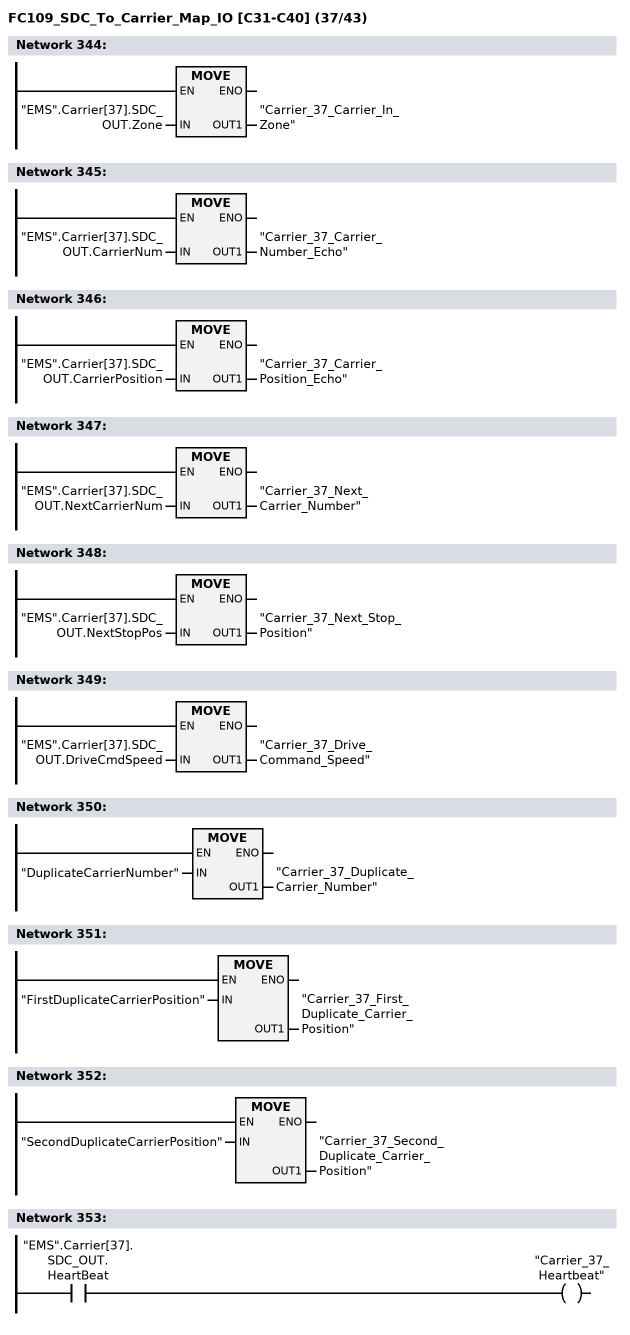
   RUNG wire#powerrail
      Move(in := "EMS".Carrier[37].SDC_OUT.Zone, out1 => "Carrier_37_Carrier_In_Zone")
   END_RUNG
   // the same network as SCL:
   "Carrier_37_Carrier_In_Zone" := "EMS".Carrier[37].SDC_OUT.Zone;
END_REGION

REGION Network 345
   RUNG wire#powerrail
      Move(in := "EMS".Carrier[37].SDC_OUT.CarrierNum, out1 => "Carrier_37_Carrier_Number_Echo")
   END_RUNG
   // the same network as SCL:
   "Carrier_37_Carrier_Number_Echo" := "EMS".Carrier[37].SDC_OUT.CarrierNum;
END_REGION

REGION Network 346
   RUNG wire#powerrail
      Move(in := "EMS".Carrier[37].SDC_OUT.CarrierPosition, out1 => "Carrier_37_Carrier_Position_Echo")
   END_RUNG
   // the same network as SCL:
   "Carrier_37_Carrier_Position_Echo" := "EMS".Carrier[37].SDC_OUT.CarrierPosition;
END_REGION

REGION Network 347
   RUNG wire#powerrail
      Move(in := "EMS".Carrier[37].SDC_OUT.NextCarrierNum, out1 => "Carrier_37_Next_Carrier_Number")
   END_RUNG
   // the same network as SCL:
   "Carrier_37_Next_Carrier_Number" := "EMS".Carrier[37].SDC_OUT.NextCarrierNum;
END_REGION

REGION Network 348
   RUNG wire#powerrail
      Move(in := "EMS".Carrier[37].SDC_OUT.NextStopPos, out1 => "Carrier_37_Next_Stop_Position")
   END_RUNG
   // the same network as SCL:
   "Carrier_37_Next_Stop_Position" := "EMS".Carrier[37].SDC_OUT.NextStopPos;
END_REGION

REGION Network 349
   RUNG wire#powerrail
      Move(in := "EMS".Carrier[37].SDC_OUT.DriveCmdSpeed, out1 => "Carrier_37_Drive_Command_Speed")
   END_RUNG
   // the same network as SCL:
   "Carrier_37_Drive_Command_Speed" := "EMS".Carrier[37].SDC_OUT.DriveCmdSpeed;
END_REGION

REGION Network 350
   RUNG wire#powerrail
      Move(in := "DuplicateCarrierNumber", out1 => "Carrier_37_Duplicate_Carrier_Number")
   END_RUNG
   // the same network as SCL:
   "Carrier_37_Duplicate_Carrier_Number" := "DuplicateCarrierNumber";
END_REGION

REGION Network 351
   RUNG wire#powerrail
      Move(in := "FirstDuplicateCarrierPosition", out1 => "Carrier_37_First_Duplicate_Carrier_Position")
   END_RUNG
   // the same network as SCL:
   "Carrier_37_First_Duplicate_Carrier_Position" := "FirstDuplicateCarrierPosition";
END_REGION

REGION Network 352
   RUNG wire#powerrail
      Move(in := "SecondDuplicateCarrierPosition", out1 => "Carrier_37_Second_Duplicate_Carrier_Position")
   END_RUNG
   // the same network as SCL:
   "Carrier_37_Second_Duplicate_Carrier_Position" := "SecondDuplicateCarrierPosition";
END_REGION

REGION Network 353
   RUNG wire#powerrail
      Contact( "EMS".Carrier[37].SDC_OUT.HeartBeat )
      Coil( "Carrier_37_Heartbeat" )
   END_RUNG
   // the same network as SCL:
   "Carrier_37_Heartbeat" := "EMS".Carrier[37].SDC_OUT.HeartBeat;
END_REGION

REGION Network 354
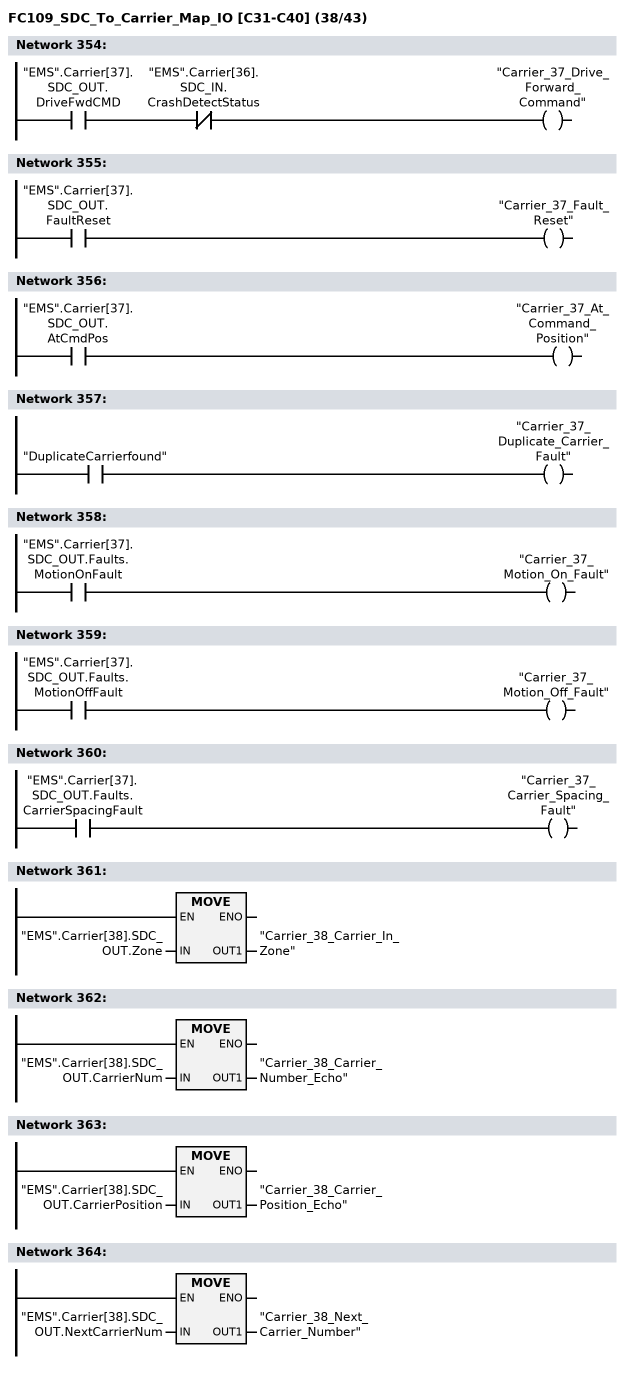
   RUNG wire#powerrail
      Contact( "EMS".Carrier[37].SDC_OUT.DriveFwdCMD )
      I_Contact( "EMS".Carrier[36].SDC_IN.CrashDetectStatus )
      Coil( "Carrier_37_Drive_Forward_Command" )
   END_RUNG
   // the same network as SCL:
   "Carrier_37_Drive_Forward_Command" := "EMS".Carrier[37].SDC_OUT.DriveFwdCMD AND NOT "EMS".Carrier[36].SDC_IN.CrashDetectStatus;
END_REGION

REGION Network 355
   RUNG wire#powerrail
      Contact( "EMS".Carrier[37].SDC_OUT.FaultReset )
      Coil( "Carrier_37_Fault_Reset" )
   END_RUNG
   // the same network as SCL:
   "Carrier_37_Fault_Reset" := "EMS".Carrier[37].SDC_OUT.FaultReset;
END_REGION

REGION Network 356
   RUNG wire#powerrail
      Contact( "EMS".Carrier[37].SDC_OUT.AtCmdPos )
      Coil( "Carrier_37_At_Command_Position" )
   END_RUNG
   // the same network as SCL:
   "Carrier_37_At_Command_Position" := "EMS".Carrier[37].SDC_OUT.AtCmdPos;
END_REGION

REGION Network 357
   RUNG wire#powerrail
      Contact( "DuplicateCarrierfound" )
      Coil( "Carrier_37_Duplicate_Carrier_Fault" )
   END_RUNG
   // the same network as SCL:
   "Carrier_37_Duplicate_Carrier_Fault" := "DuplicateCarrierfound";
END_REGION

REGION Network 358
   RUNG wire#powerrail
      Contact( "EMS".Carrier[37].SDC_OUT.Faults.MotionOnFault )
      Coil( "Carrier_37_Motion_On_Fault" )
   END_RUNG
   // the same network as SCL:
   "Carrier_37_Motion_On_Fault" := "EMS".Carrier[37].SDC_OUT.Faults.MotionOnFault;
END_REGION

REGION Network 359
   RUNG wire#powerrail
      Contact( "EMS".Carrier[37].SDC_OUT.Faults.MotionOffFault )
      Coil( "Carrier_37_Motion_Off_Fault" )
   END_RUNG
   // the same network as SCL:
   "Carrier_37_Motion_Off_Fault" := "EMS".Carrier[37].SDC_OUT.Faults.MotionOffFault;
END_REGION

REGION Network 360
   RUNG wire#powerrail
      Contact( "EMS".Carrier[37].SDC_OUT.Faults.CarrierSpacingFault )
      Coil( "Carrier_37_Carrier_Spacing_Fault" )
   END_RUNG
   // the same network as SCL:
   "Carrier_37_Carrier_Spacing_Fault" := "EMS".Carrier[37].SDC_OUT.Faults.CarrierSpacingFault;
END_REGION

REGION Network 361
   RUNG wire#powerrail
      Move(in := "EMS".Carrier[38].SDC_OUT.Zone, out1 => "Carrier_38_Carrier_In_Zone")
   END_RUNG
   // the same network as SCL:
   "Carrier_38_Carrier_In_Zone" := "EMS".Carrier[38].SDC_OUT.Zone;
END_REGION

REGION Network 362
   RUNG wire#powerrail
      Move(in := "EMS".Carrier[38].SDC_OUT.CarrierNum, out1 => "Carrier_38_Carrier_Number_Echo")
   END_RUNG
   // the same network as SCL:
   "Carrier_38_Carrier_Number_Echo" := "EMS".Carrier[38].SDC_OUT.CarrierNum;
END_REGION

REGION Network 363
   RUNG wire#powerrail
      Move(in := "EMS".Carrier[38].SDC_OUT.CarrierPosition, out1 => "Carrier_38_Carrier_Position_Echo")
   END_RUNG
   // the same network as SCL:
   "Carrier_38_Carrier_Position_Echo" := "EMS".Carrier[38].SDC_OUT.CarrierPosition;
END_REGION

REGION Network 364
   RUNG wire#powerrail
      Move(in := "EMS".Carrier[38].SDC_OUT.NextCarrierNum, out1 => "Carrier_38_Next_Carrier_Number")
   END_RUNG
   // the same network as SCL:
   "Carrier_38_Next_Carrier_Number" := "EMS".Carrier[38].SDC_OUT.NextCarrierNum;
END_REGION

REGION Network 365
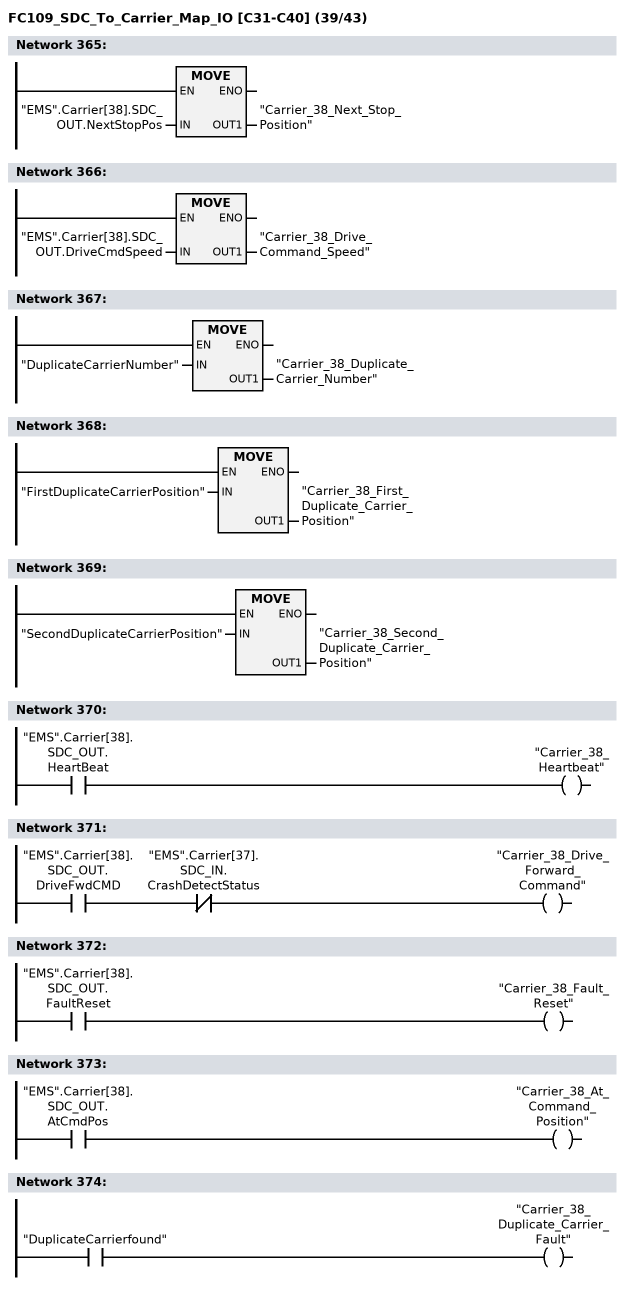
   RUNG wire#powerrail
      Move(in := "EMS".Carrier[38].SDC_OUT.NextStopPos, out1 => "Carrier_38_Next_Stop_Position")
   END_RUNG
   // the same network as SCL:
   "Carrier_38_Next_Stop_Position" := "EMS".Carrier[38].SDC_OUT.NextStopPos;
END_REGION

REGION Network 366
   RUNG wire#powerrail
      Move(in := "EMS".Carrier[38].SDC_OUT.DriveCmdSpeed, out1 => "Carrier_38_Drive_Command_Speed")
   END_RUNG
   // the same network as SCL:
   "Carrier_38_Drive_Command_Speed" := "EMS".Carrier[38].SDC_OUT.DriveCmdSpeed;
END_REGION

REGION Network 367
   RUNG wire#powerrail
      Move(in := "DuplicateCarrierNumber", out1 => "Carrier_38_Duplicate_Carrier_Number")
   END_RUNG
   // the same network as SCL:
   "Carrier_38_Duplicate_Carrier_Number" := "DuplicateCarrierNumber";
END_REGION

REGION Network 368
   RUNG wire#powerrail
      Move(in := "FirstDuplicateCarrierPosition", out1 => "Carrier_38_First_Duplicate_Carrier_Position")
   END_RUNG
   // the same network as SCL:
   "Carrier_38_First_Duplicate_Carrier_Position" := "FirstDuplicateCarrierPosition";
END_REGION

REGION Network 369
   RUNG wire#powerrail
      Move(in := "SecondDuplicateCarrierPosition", out1 => "Carrier_38_Second_Duplicate_Carrier_Position")
   END_RUNG
   // the same network as SCL:
   "Carrier_38_Second_Duplicate_Carrier_Position" := "SecondDuplicateCarrierPosition";
END_REGION

REGION Network 370
   RUNG wire#powerrail
      Contact( "EMS".Carrier[38].SDC_OUT.HeartBeat )
      Coil( "Carrier_38_Heartbeat" )
   END_RUNG
   // the same network as SCL:
   "Carrier_38_Heartbeat" := "EMS".Carrier[38].SDC_OUT.HeartBeat;
END_REGION

REGION Network 371
   RUNG wire#powerrail
      Contact( "EMS".Carrier[38].SDC_OUT.DriveFwdCMD )
      I_Contact( "EMS".Carrier[37].SDC_IN.CrashDetectStatus )
      Coil( "Carrier_38_Drive_Forward_Command" )
   END_RUNG
   // the same network as SCL:
   "Carrier_38_Drive_Forward_Command" := "EMS".Carrier[38].SDC_OUT.DriveFwdCMD AND NOT "EMS".Carrier[37].SDC_IN.CrashDetectStatus;
END_REGION

REGION Network 372
   RUNG wire#powerrail
      Contact( "EMS".Carrier[38].SDC_OUT.FaultReset )
      Coil( "Carrier_38_Fault_Reset" )
   END_RUNG
   // the same network as SCL:
   "Carrier_38_Fault_Reset" := "EMS".Carrier[38].SDC_OUT.FaultReset;
END_REGION

REGION Network 373
   RUNG wire#powerrail
      Contact( "EMS".Carrier[38].SDC_OUT.AtCmdPos )
      Coil( "Carrier_38_At_Command_Position" )
   END_RUNG
   // the same network as SCL:
   "Carrier_38_At_Command_Position" := "EMS".Carrier[38].SDC_OUT.AtCmdPos;
END_REGION

REGION Network 374
   RUNG wire#powerrail
      Contact( "DuplicateCarrierfound" )
      Coil( "Carrier_38_Duplicate_Carrier_Fault" )
   END_RUNG
   // the same network as SCL:
   "Carrier_38_Duplicate_Carrier_Fault" := "DuplicateCarrierfound";
END_REGION

REGION Network 375
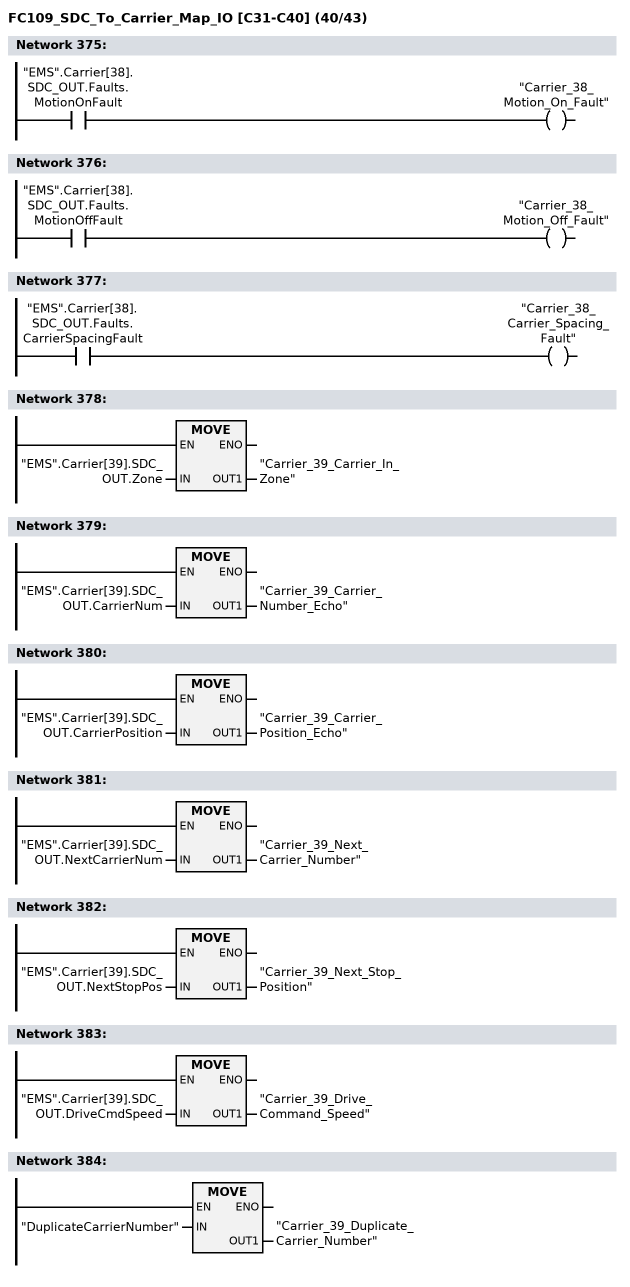
   RUNG wire#powerrail
      Contact( "EMS".Carrier[38].SDC_OUT.Faults.MotionOnFault )
      Coil( "Carrier_38_Motion_On_Fault" )
   END_RUNG
   // the same network as SCL:
   "Carrier_38_Motion_On_Fault" := "EMS".Carrier[38].SDC_OUT.Faults.MotionOnFault;
END_REGION

REGION Network 376
   RUNG wire#powerrail
      Contact( "EMS".Carrier[38].SDC_OUT.Faults.MotionOffFault )
      Coil( "Carrier_38_Motion_Off_Fault" )
   END_RUNG
   // the same network as SCL:
   "Carrier_38_Motion_Off_Fault" := "EMS".Carrier[38].SDC_OUT.Faults.MotionOffFault;
END_REGION

REGION Network 377
   RUNG wire#powerrail
      Contact( "EMS".Carrier[38].SDC_OUT.Faults.CarrierSpacingFault )
      Coil( "Carrier_38_Carrier_Spacing_Fault" )
   END_RUNG
   // the same network as SCL:
   "Carrier_38_Carrier_Spacing_Fault" := "EMS".Carrier[38].SDC_OUT.Faults.CarrierSpacingFault;
END_REGION

REGION Network 378
   RUNG wire#powerrail
      Move(in := "EMS".Carrier[39].SDC_OUT.Zone, out1 => "Carrier_39_Carrier_In_Zone")
   END_RUNG
   // the same network as SCL:
   "Carrier_39_Carrier_In_Zone" := "EMS".Carrier[39].SDC_OUT.Zone;
END_REGION

REGION Network 379
   RUNG wire#powerrail
      Move(in := "EMS".Carrier[39].SDC_OUT.CarrierNum, out1 => "Carrier_39_Carrier_Number_Echo")
   END_RUNG
   // the same network as SCL:
   "Carrier_39_Carrier_Number_Echo" := "EMS".Carrier[39].SDC_OUT.CarrierNum;
END_REGION

REGION Network 380
   RUNG wire#powerrail
      Move(in := "EMS".Carrier[39].SDC_OUT.CarrierPosition, out1 => "Carrier_39_Carrier_Position_Echo")
   END_RUNG
   // the same network as SCL:
   "Carrier_39_Carrier_Position_Echo" := "EMS".Carrier[39].SDC_OUT.CarrierPosition;
END_REGION

REGION Network 381
   RUNG wire#powerrail
      Move(in := "EMS".Carrier[39].SDC_OUT.NextCarrierNum, out1 => "Carrier_39_Next_Carrier_Number")
   END_RUNG
   // the same network as SCL:
   "Carrier_39_Next_Carrier_Number" := "EMS".Carrier[39].SDC_OUT.NextCarrierNum;
END_REGION

REGION Network 382
   RUNG wire#powerrail
      Move(in := "EMS".Carrier[39].SDC_OUT.NextStopPos, out1 => "Carrier_39_Next_Stop_Position")
   END_RUNG
   // the same network as SCL:
   "Carrier_39_Next_Stop_Position" := "EMS".Carrier[39].SDC_OUT.NextStopPos;
END_REGION

REGION Network 383
   RUNG wire#powerrail
      Move(in := "EMS".Carrier[39].SDC_OUT.DriveCmdSpeed, out1 => "Carrier_39_Drive_Command_Speed")
   END_RUNG
   // the same network as SCL:
   "Carrier_39_Drive_Command_Speed" := "EMS".Carrier[39].SDC_OUT.DriveCmdSpeed;
END_REGION

REGION Network 384
   RUNG wire#powerrail
      Move(in := "DuplicateCarrierNumber", out1 => "Carrier_39_Duplicate_Carrier_Number")
   END_RUNG
   // the same network as SCL:
   "Carrier_39_Duplicate_Carrier_Number" := "DuplicateCarrierNumber";
END_REGION

REGION Network 385
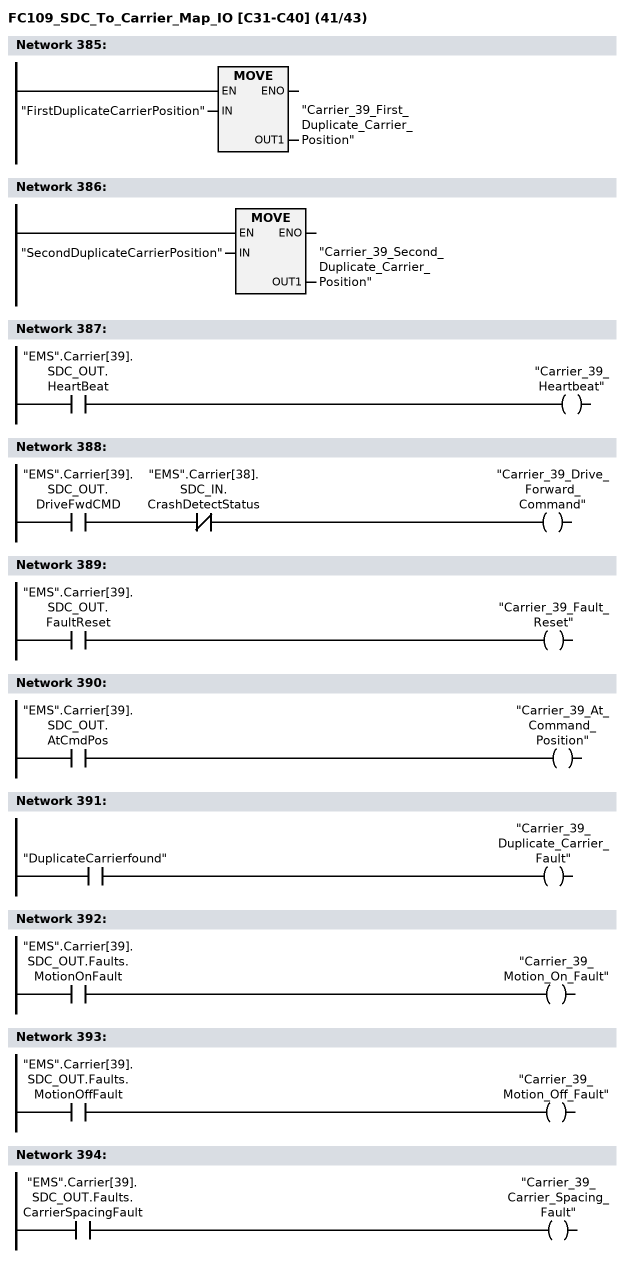
   RUNG wire#powerrail
      Move(in := "FirstDuplicateCarrierPosition", out1 => "Carrier_39_First_Duplicate_Carrier_Position")
   END_RUNG
   // the same network as SCL:
   "Carrier_39_First_Duplicate_Carrier_Position" := "FirstDuplicateCarrierPosition";
END_REGION

REGION Network 386
   RUNG wire#powerrail
      Move(in := "SecondDuplicateCarrierPosition", out1 => "Carrier_39_Second_Duplicate_Carrier_Position")
   END_RUNG
   // the same network as SCL:
   "Carrier_39_Second_Duplicate_Carrier_Position" := "SecondDuplicateCarrierPosition";
END_REGION

REGION Network 387
   RUNG wire#powerrail
      Contact( "EMS".Carrier[39].SDC_OUT.HeartBeat )
      Coil( "Carrier_39_Heartbeat" )
   END_RUNG
   // the same network as SCL:
   "Carrier_39_Heartbeat" := "EMS".Carrier[39].SDC_OUT.HeartBeat;
END_REGION

REGION Network 388
   RUNG wire#powerrail
      Contact( "EMS".Carrier[39].SDC_OUT.DriveFwdCMD )
      I_Contact( "EMS".Carrier[38].SDC_IN.CrashDetectStatus )
      Coil( "Carrier_39_Drive_Forward_Command" )
   END_RUNG
   // the same network as SCL:
   "Carrier_39_Drive_Forward_Command" := "EMS".Carrier[39].SDC_OUT.DriveFwdCMD AND NOT "EMS".Carrier[38].SDC_IN.CrashDetectStatus;
END_REGION

REGION Network 389
   RUNG wire#powerrail
      Contact( "EMS".Carrier[39].SDC_OUT.FaultReset )
      Coil( "Carrier_39_Fault_Reset" )
   END_RUNG
   // the same network as SCL:
   "Carrier_39_Fault_Reset" := "EMS".Carrier[39].SDC_OUT.FaultReset;
END_REGION

REGION Network 390
   RUNG wire#powerrail
      Contact( "EMS".Carrier[39].SDC_OUT.AtCmdPos )
      Coil( "Carrier_39_At_Command_Position" )
   END_RUNG
   // the same network as SCL:
   "Carrier_39_At_Command_Position" := "EMS".Carrier[39].SDC_OUT.AtCmdPos;
END_REGION

REGION Network 391
   RUNG wire#powerrail
      Contact( "DuplicateCarrierfound" )
      Coil( "Carrier_39_Duplicate_Carrier_Fault" )
   END_RUNG
   // the same network as SCL:
   "Carrier_39_Duplicate_Carrier_Fault" := "DuplicateCarrierfound";
END_REGION

REGION Network 392
   RUNG wire#powerrail
      Contact( "EMS".Carrier[39].SDC_OUT.Faults.MotionOnFault )
      Coil( "Carrier_39_Motion_On_Fault" )
   END_RUNG
   // the same network as SCL:
   "Carrier_39_Motion_On_Fault" := "EMS".Carrier[39].SDC_OUT.Faults.MotionOnFault;
END_REGION

REGION Network 393
   RUNG wire#powerrail
      Contact( "EMS".Carrier[39].SDC_OUT.Faults.MotionOffFault )
      Coil( "Carrier_39_Motion_Off_Fault" )
   END_RUNG
   // the same network as SCL:
   "Carrier_39_Motion_Off_Fault" := "EMS".Carrier[39].SDC_OUT.Faults.MotionOffFault;
END_REGION

REGION Network 394
   RUNG wire#powerrail
      Contact( "EMS".Carrier[39].SDC_OUT.Faults.CarrierSpacingFault )
      Coil( "Carrier_39_Carrier_Spacing_Fault" )
   END_RUNG
   // the same network as SCL:
   "Carrier_39_Carrier_Spacing_Fault" := "EMS".Carrier[39].SDC_OUT.Faults.CarrierSpacingFault;
END_REGION

REGION Network 395
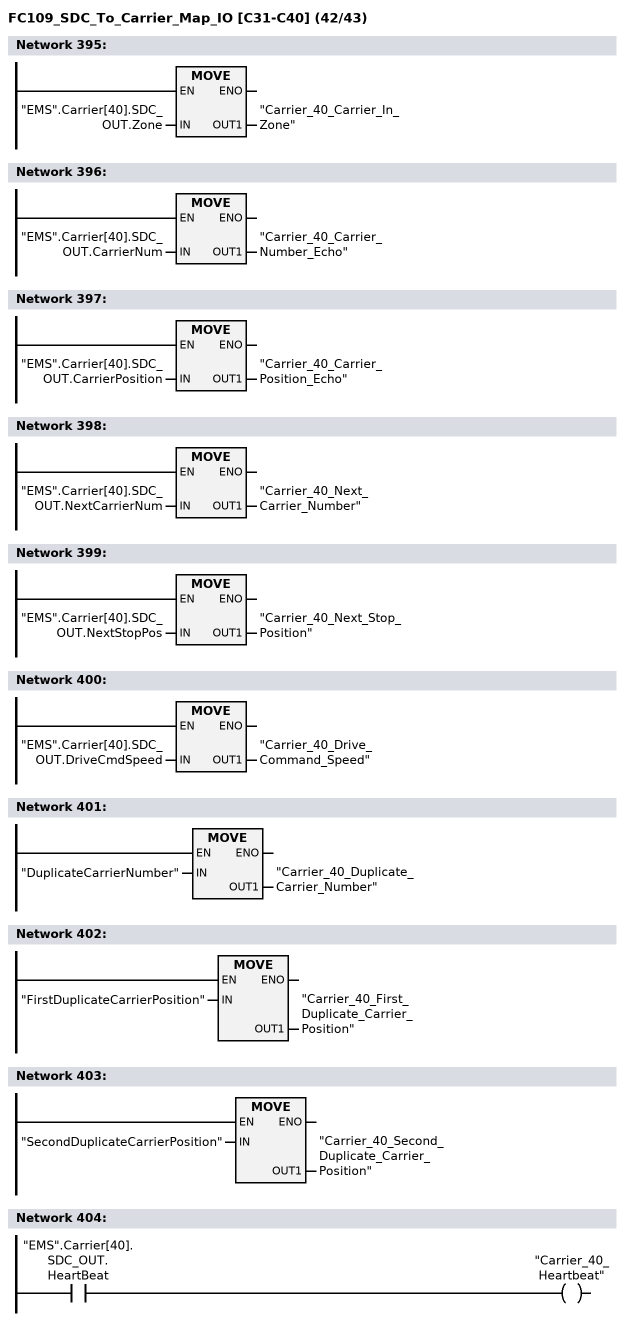
   RUNG wire#powerrail
      Move(in := "EMS".Carrier[40].SDC_OUT.Zone, out1 => "Carrier_40_Carrier_In_Zone")
   END_RUNG
   // the same network as SCL:
   "Carrier_40_Carrier_In_Zone" := "EMS".Carrier[40].SDC_OUT.Zone;
END_REGION

REGION Network 396
   RUNG wire#powerrail
      Move(in := "EMS".Carrier[40].SDC_OUT.CarrierNum, out1 => "Carrier_40_Carrier_Number_Echo")
   END_RUNG
   // the same network as SCL:
   "Carrier_40_Carrier_Number_Echo" := "EMS".Carrier[40].SDC_OUT.CarrierNum;
END_REGION

REGION Network 397
   RUNG wire#powerrail
      Move(in := "EMS".Carrier[40].SDC_OUT.CarrierPosition, out1 => "Carrier_40_Carrier_Position_Echo")
   END_RUNG
   // the same network as SCL:
   "Carrier_40_Carrier_Position_Echo" := "EMS".Carrier[40].SDC_OUT.CarrierPosition;
END_REGION

REGION Network 398
   RUNG wire#powerrail
      Move(in := "EMS".Carrier[40].SDC_OUT.NextCarrierNum, out1 => "Carrier_40_Next_Carrier_Number")
   END_RUNG
   // the same network as SCL:
   "Carrier_40_Next_Carrier_Number" := "EMS".Carrier[40].SDC_OUT.NextCarrierNum;
END_REGION

REGION Network 399
   RUNG wire#powerrail
      Move(in := "EMS".Carrier[40].SDC_OUT.NextStopPos, out1 => "Carrier_40_Next_Stop_Position")
   END_RUNG
   // the same network as SCL:
   "Carrier_40_Next_Stop_Position" := "EMS".Carrier[40].SDC_OUT.NextStopPos;
END_REGION

REGION Network 400
   RUNG wire#powerrail
      Move(in := "EMS".Carrier[40].SDC_OUT.DriveCmdSpeed, out1 => "Carrier_40_Drive_Command_Speed")
   END_RUNG
   // the same network as SCL:
   "Carrier_40_Drive_Command_Speed" := "EMS".Carrier[40].SDC_OUT.DriveCmdSpeed;
END_REGION

REGION Network 401
   RUNG wire#powerrail
      Move(in := "DuplicateCarrierNumber", out1 => "Carrier_40_Duplicate_Carrier_Number")
   END_RUNG
   // the same network as SCL:
   "Carrier_40_Duplicate_Carrier_Number" := "DuplicateCarrierNumber";
END_REGION

REGION Network 402
   RUNG wire#powerrail
      Move(in := "FirstDuplicateCarrierPosition", out1 => "Carrier_40_First_Duplicate_Carrier_Position")
   END_RUNG
   // the same network as SCL:
   "Carrier_40_First_Duplicate_Carrier_Position" := "FirstDuplicateCarrierPosition";
END_REGION

REGION Network 403
   RUNG wire#powerrail
      Move(in := "SecondDuplicateCarrierPosition", out1 => "Carrier_40_Second_Duplicate_Carrier_Position")
   END_RUNG
   // the same network as SCL:
   "Carrier_40_Second_Duplicate_Carrier_Position" := "SecondDuplicateCarrierPosition";
END_REGION

REGION Network 404
   RUNG wire#powerrail
      Contact( "EMS".Carrier[40].SDC_OUT.HeartBeat )
      Coil( "Carrier_40_Heartbeat" )
   END_RUNG
   // the same network as SCL:
   "Carrier_40_Heartbeat" := "EMS".Carrier[40].SDC_OUT.HeartBeat;
END_REGION

REGION Network 405
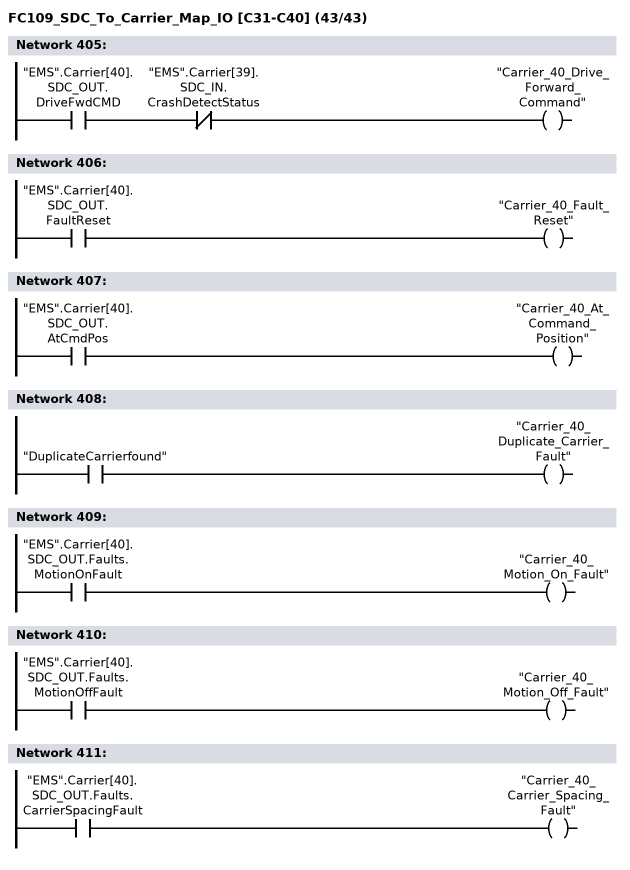
   RUNG wire#powerrail
      Contact( "EMS".Carrier[40].SDC_OUT.DriveFwdCMD )
      I_Contact( "EMS".Carrier[39].SDC_IN.CrashDetectStatus )
      Coil( "Carrier_40_Drive_Forward_Command" )
   END_RUNG
   // the same network as SCL:
   "Carrier_40_Drive_Forward_Command" := "EMS".Carrier[40].SDC_OUT.DriveFwdCMD AND NOT "EMS".Carrier[39].SDC_IN.CrashDetectStatus;
END_REGION

REGION Network 406
   RUNG wire#powerrail
      Contact( "EMS".Carrier[40].SDC_OUT.FaultReset )
      Coil( "Carrier_40_Fault_Reset" )
   END_RUNG
   // the same network as SCL:
   "Carrier_40_Fault_Reset" := "EMS".Carrier[40].SDC_OUT.FaultReset;
END_REGION

REGION Network 407
   RUNG wire#powerrail
      Contact( "EMS".Carrier[40].SDC_OUT.AtCmdPos )
      Coil( "Carrier_40_At_Command_Position" )
   END_RUNG
   // the same network as SCL:
   "Carrier_40_At_Command_Position" := "EMS".Carrier[40].SDC_OUT.AtCmdPos;
END_REGION

REGION Network 408
   RUNG wire#powerrail
      Contact( "DuplicateCarrierfound" )
      Coil( "Carrier_40_Duplicate_Carrier_Fault" )
   END_RUNG
   // the same network as SCL:
   "Carrier_40_Duplicate_Carrier_Fault" := "DuplicateCarrierfound";
END_REGION

REGION Network 409
   RUNG wire#powerrail
      Contact( "EMS".Carrier[40].SDC_OUT.Faults.MotionOnFault )
      Coil( "Carrier_40_Motion_On_Fault" )
   END_RUNG
   // the same network as SCL:
   "Carrier_40_Motion_On_Fault" := "EMS".Carrier[40].SDC_OUT.Faults.MotionOnFault;
END_REGION

REGION Network 410
   RUNG wire#powerrail
      Contact( "EMS".Carrier[40].SDC_OUT.Faults.MotionOffFault )
      Coil( "Carrier_40_Motion_Off_Fault" )
   END_RUNG
   // the same network as SCL:
   "Carrier_40_Motion_Off_Fault" := "EMS".Carrier[40].SDC_OUT.Faults.MotionOffFault;
END_REGION

REGION Network 411
   RUNG wire#powerrail
      Contact( "EMS".Carrier[40].SDC_OUT.Faults.CarrierSpacingFault )
      Coil( "Carrier_40_Carrier_Spacing_Fault" )
   END_RUNG
   // the same network as SCL:
   "Carrier_40_Carrier_Spacing_Fault" := "EMS".Carrier[40].SDC_OUT.Faults.CarrierSpacingFault;
END_REGION
END_FUNCTION

FUNCTION "FC110_SDC_To_Carrier_Map_IO [C41-C50]" : Void   // FC110, LAD
{ S7_Optimized_Access := 'TRUE' }
VERSION : 0.1
BEGIN

REGION Network 1
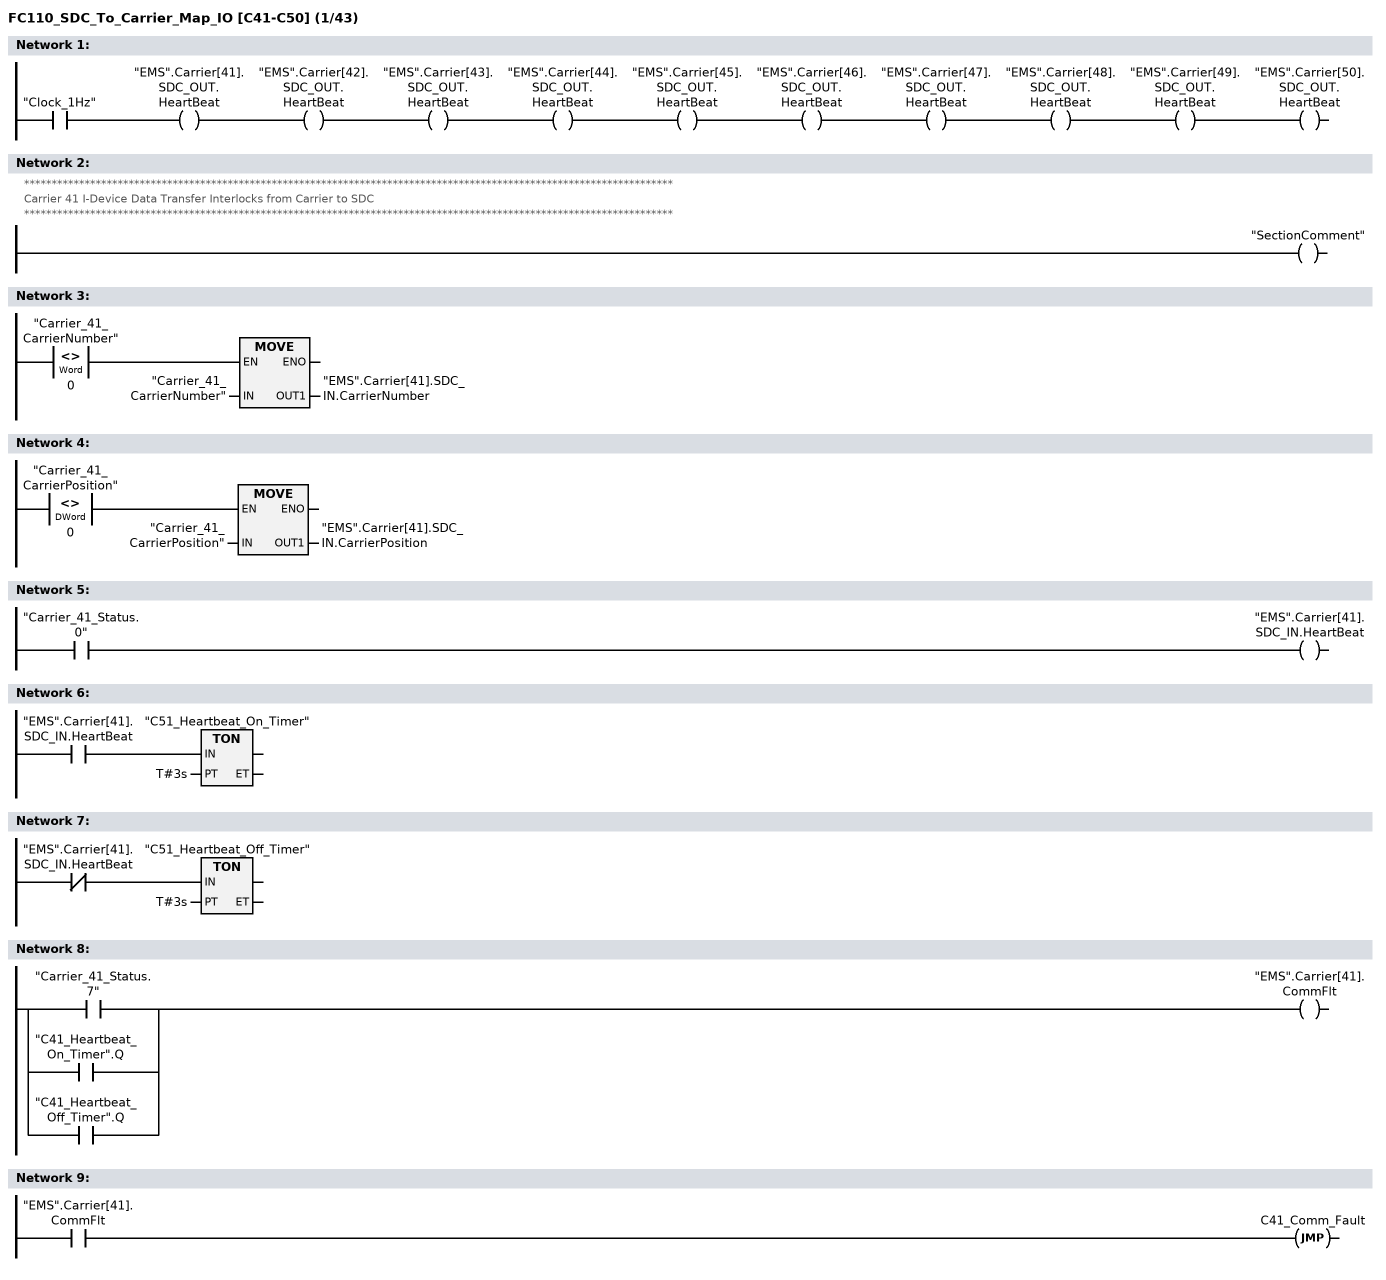
   RUNG wire#powerrail
      Contact( "Clock_1Hz" )
      Coil( "EMS".Carrier[41].SDC_OUT.HeartBeat )
      Coil( "EMS".Carrier[42].SDC_OUT.HeartBeat )
      Coil( "EMS".Carrier[43].SDC_OUT.HeartBeat )
      Coil( "EMS".Carrier[44].SDC_OUT.HeartBeat )
      Coil( "EMS".Carrier[45].SDC_OUT.HeartBeat )
      Coil( "EMS".Carrier[46].SDC_OUT.HeartBeat )
      Coil( "EMS".Carrier[47].SDC_OUT.HeartBeat )
      Coil( "EMS".Carrier[48].SDC_OUT.HeartBeat )
      Coil( "EMS".Carrier[49].SDC_OUT.HeartBeat )
      Coil( "EMS".Carrier[50].SDC_OUT.HeartBeat )
   END_RUNG
   // the same network as SCL:
   "EMS".Carrier[41].SDC_OUT.HeartBeat := "Clock_1Hz";
   "EMS".Carrier[42].SDC_OUT.HeartBeat := "Clock_1Hz";
   "EMS".Carrier[43].SDC_OUT.HeartBeat := "Clock_1Hz";
   "EMS".Carrier[44].SDC_OUT.HeartBeat := "Clock_1Hz";
   "EMS".Carrier[45].SDC_OUT.HeartBeat := "Clock_1Hz";
   "EMS".Carrier[46].SDC_OUT.HeartBeat := "Clock_1Hz";
   "EMS".Carrier[47].SDC_OUT.HeartBeat := "Clock_1Hz";
   "EMS".Carrier[48].SDC_OUT.HeartBeat := "Clock_1Hz";
   "EMS".Carrier[49].SDC_OUT.HeartBeat := "Clock_1Hz";
   "EMS".Carrier[50].SDC_OUT.HeartBeat := "Clock_1Hz";
END_REGION

REGION Network 2
   // **********************************************************************************************************************
   // 
   // Carrier 41 I-Device Data Transfer Interlocks from Carrier to SDC
   // 
   // **********************************************************************************************************************
   RUNG wire#powerrail
      Coil( "SectionComment" )
   END_RUNG
   // the same network as SCL:
   "SectionComment" := TRUE;
END_REGION

REGION Network 3
   RUNG wire#powerrail
      { S7_Templates := "SrcType := Word" } NE_Contact(in1 := "Carrier_41_CarrierNumber", in2 := 0)
      Move(in := "Carrier_41_CarrierNumber", out1 => "EMS".Carrier[41].SDC_IN.CarrierNumber)
   END_RUNG
   // the same network as SCL:
   IF "Carrier_41_CarrierNumber" <> 0 THEN
       "EMS".Carrier[41].SDC_IN.CarrierNumber := "Carrier_41_CarrierNumber";
   END_IF;
END_REGION

REGION Network 4
   RUNG wire#powerrail
      { S7_Templates := "SrcType := DWord" } NE_Contact(in1 := "Carrier_41_CarrierPosition", in2 := 0)
      Move(in := "Carrier_41_CarrierPosition", out1 => "EMS".Carrier[41].SDC_IN.CarrierPosition)
   END_RUNG
   // the same network as SCL:
   IF "Carrier_41_CarrierPosition" <> 0 THEN
       "EMS".Carrier[41].SDC_IN.CarrierPosition := "Carrier_41_CarrierPosition";
   END_IF;
END_REGION

REGION Network 5
   RUNG wire#powerrail
      Contact( "Carrier_41_Status.0" )
      Coil( "EMS".Carrier[41].SDC_IN.HeartBeat )
   END_RUNG
   // the same network as SCL:
   "EMS".Carrier[41].SDC_IN.HeartBeat := "Carrier_41_Status.0";
END_REGION

REGION Network 6
   "C51_Heartbeat_On_Timer".TON(IN := "EMS".Carrier[41].SDC_IN.HeartBeat, PT := T#3s);
END_REGION

REGION Network 7
   "C51_Heartbeat_Off_Timer".TON(IN := NOT "EMS".Carrier[41].SDC_IN.HeartBeat, PT := T#3s);
END_REGION

REGION Network 8
   RUNG wire#powerrail
      Contact( "Carrier_41_Status.7" )
      wire#w1
      Coil( "EMS".Carrier[41].CommFlt )
   END_RUNG
   RUNG wire#powerrail
      Contact( "C41_Heartbeat_On_Timer".Q )
   END_RUNG wire#w1
   RUNG wire#powerrail
      Contact( "C41_Heartbeat_Off_Timer".Q )
   END_RUNG wire#w1
   // the same network as SCL:
   "EMS".Carrier[41].CommFlt := "Carrier_41_Status.7" OR "C41_Heartbeat_On_Timer".Q OR "C41_Heartbeat_Off_Timer".Q;
END_REGION

REGION Network 9
   RUNG wire#powerrail
      Contact( "EMS".Carrier[41].CommFlt )
      JumpCoil( C41_Comm_Fault )
   END_RUNG
   // the same network as SCL:
   IF "EMS".Carrier[41].CommFlt THEN GOTO C41_Comm_Fault; END_IF;
END_REGION

REGION Network 10